PopupScreen "Tank 6S Status" 480x272
   TextField "Text field_4" at 9,135 size 86x22; Text 'Pressure:'
   IOField "I/O field_1" at 148,130 size 90x25; FormatPattern s999.9; Unit  mBar
      ProcessValue <- "20_TANKS_IP_DATA_RIO_06_SECOND_TANK_TANKS_PRESS"
   TextField "Text field_5" at 9,169 size 113x22; Text 'Water Level:'
   IOField "I/O field_2" at 148,164 size 90x25; FormatPattern 999.9; Unit  %
      ProcessValue <- "20_TANKS_IP_DATA_RIO_06_SECOND_TANK_BWT_LEVEL"
   TextField "Text field_6" at 9,203 size 137x22; Text 'MBG Flow Rate:'
   IOField "I/O field_3" at 148,198 size 90x25; FormatPattern 999.9; Unit  m³/hr
      ProcessValue <- "20_TANKS_IP_DATA_RIO_06_SECOND_TANK_MBG_FLOW"
   TextField "Text field_7" at 9,237 size 135x22; Text 'USD Flow Rate:'
   IOField "I/O field_4" at 148,232 size 90x25; FormatPattern 999.9; Unit  m³/hr
      ProcessValue <- "20_TANKS_IP_DATA_RIO_06_SECOND_TANK_USD_FLOW"
   Button "Button_1" at 51,5 size 191x35; TextOff 'Starboard Tank 6 (6S)'
      on Release: function_efd93a16("Tank 6S Status", 0, 0, -1, 2, 1)
   TextField "Text field_1" at 6,90 size 109x25; Text 'TIME LEFT:'
   GraphicView "Graphic view_1" at 9,46 size 228x32; Picture "Tank Manually Disabled"
   GraphicIOField "Graphic I/O field_1" at 9,46 size 228x32; PictureList "Tank Process Stage_II"
      ProcessValue <- "2100_BTCS_CNTRL_DB_BTCS_STATE"
      Visibility <- "504_Tank Grouping_DB2020_GROUP of TANK 13"
   Button "Button_2" at 4,5 size 45x35; TextOff 'Text'; PictureOff "Graphic_286"
      on Click: function_efd93a16("Tank 6S Status", 0, 0, -1, -1, 1)
   IOField "I/O field_29" at 190,90 size 47x25; FormatPattern 99; Unit m
      ProcessValue <- "504_Tank Grouping_DB2020_Time Left Tank_Time Left m Tank 13"
   IOField "I/O field_8" at 147,90 size 42x25; FormatPattern 99; Unit h
      ProcessValue <- "504_Tank Grouping_DB2020_Time Left Tank_Time Left h Tank 13"
   IOField "I/O field_9" at 104,90 size 42x25; FormatPattern 99; Unit d
      ProcessValue <- "504_Tank Grouping_DB2020_Time Left Tank_Time Left d Tank 13"
   TextField "Text field_8" at 244,135 size 140x22; Text 'Water pH Level:'
   IOField "I/O field_5" at 384,130 size 90x25; FormatPattern 99.9
      ProcessValue <- "20_TANKS_IP_DATA_RIO_06_SECOND_TANK_BWT_PH"
   TextField "Text field_9" at 244,169 size 143x22; Text 'Water DO Level:'
   IOField "I/O field_6" at 384,164 size 90x25; FormatPattern 99.99; Unit  mg/l
      ProcessValue <- "20_TANKS_IP_DATA_RIO_06_SECOND_TANK_BWT_DO"
   TextField "Text field_10" at 244,203 size 174x22; Text 'Water Temperature:'
   IOField "I/O field_7" at 399,198 size 75x25; FormatPattern 999.9; Unit  °C
      ProcessValue <- "20_TANKS_IP_DATA_RIO_06_SECOND_TANK_BWT_TEMP"
   Group "Group" at 248,228 size 226x40
   Button "Button_5" at 248,228 size 226x40; TextOff 'Tank Shutdown Alarm'
      Visibility <- "2062_Warning_Data_Alarm Tank S6"
   Button "Button_6" at 248,228 size 226x40; TextOff 'No/Low Water Level'; Authorization "Operate"
      Visibility <- "LT421 6S  TANK LEVEL ALARM_ALARM L"

PopupScreen "Tank 6P Status" 480x272
   TextField "Text field_4" at 9,135 size 86x22; Text 'Pressure:'
   IOField "I/O field_1" at 147,130 size 90x25; FormatPattern s999.9; Unit  mBar
      ProcessValue <- "20_TANKS_IP_DATA_RIO_06_FIRST_TANK_TANKS_PRESS"
   TextField "Text field_5" at 9,169 size 113x22; Text 'Water Level:'
   IOField "I/O field_2" at 147,164 size 90x25; FormatPattern 999.9; Unit  %
      ProcessValue <- "20_TANKS_IP_DATA_RIO_06_FIRST_TANK_BWT_LEVEL"
   TextField "Text field_6" at 9,203 size 137x22; Text 'MBG Flow Rate:'
   IOField "I/O field_3" at 147,198 size 90x25; FormatPattern 999.9; Unit  m³/hr
      ProcessValue <- "20_TANKS_IP_DATA_RIO_06_FIRST_TANK_MBG_FLOW"
   TextField "Text field_7" at 9,237 size 135x22; Text 'USD Flow Rate:'
   IOField "I/O field_4" at 147,232 size 90x25; FormatPattern 999.9; Unit  m³/hr
      ProcessValue <- "20_TANKS_IP_DATA_RIO_06_FIRST_TANK_USD_FLOW"
   Button "Button_1" at 51,5 size 190x35; TextOff 'Port Tank 6 (6P)'
      on Release: function_efd93a16("Tank 6P Status", 0, 0, -1, 2, 1)
   TextField "Text field_1" at 5,90 size 109x25; Text 'TIME LEFT:'
   GraphicView "Graphic view_1" at 9,46 size 227x32; Picture "Tank Manually Disabled"
   GraphicIOField "Graphic I/O field_1" at 9,46 size 227x32; PictureList "Tank Process Stage_II"
      ProcessValue <- "2100_BTCS_CNTRL_DB_BTCS_STATE"
      Visibility <- "504_Tank Grouping_DB2020_GROUP of TANK 12"
   Button "Button_2" at 4,5 size 45x35; TextOff 'Text'; PictureOff "Graphic_286"
      on Click: function_efd93a16("Tank 6P Status", 0, 0, -1, -1, 1)
   IOField "I/O field_29" at 189,90 size 47x25; FormatPattern 99; Unit m
      ProcessValue <- "504_Tank Grouping_DB2020_Time Left Tank_Time Left m Tank 12"
   IOField "I/O field_8" at 146,90 size 42x25; FormatPattern 99; Unit h
      ProcessValue <- "504_Tank Grouping_DB2020_Time Left Tank_Time Left h Tank 12"
   IOField "I/O field_9" at 103,90 size 42x25; FormatPattern 99; Unit d
      ProcessValue <- "504_Tank Grouping_DB2020_Time Left Tank_Time Left d Tank 12"
   TextField "Text field_8" at 242,135 size 140x22; Text 'Water pH Level:'
   IOField "I/O field_5" at 381,130 size 90x25; FormatPattern 99.9
      ProcessValue <- "20_TANKS_IP_DATA_RIO_06_FIRST_TANK_BWT_PH"
   TextField "Text field_9" at 242,169 size 143x22; Text 'Water DO Level:'
   IOField "I/O field_6" at 381,164 size 90x25; FormatPattern 99.99; Unit  mg/l
      ProcessValue <- "20_TANKS_IP_DATA_RIO_06_FIRST_TANK_BWT_DO"
   TextField "Text field_10" at 242,203 size 174x22; Text 'Water Temperature:'
   IOField "I/O field_7" at 396,198 size 75x25; FormatPattern 999.9; Unit  °C
      ProcessValue <- "20_TANKS_IP_DATA_RIO_06_FIRST_TANK_BWT_TEMP"
   Group "Group" at 245,227 size 226x40
   Button "Button_5" at 245,227 size 226x40; TextOff 'Tank Shutdown Alarm'
      Visibility <- "2062_Warning_Data_Alarm Tank P6"
   Button "Button_6" at 245,227 size 226x40; TextOff 'No/Low Water Level'; Authorization "Operate"
      Visibility <- "LT422 6P  TANK LEVEL ALARM_ALARM L"

PopupScreen "Tank AP Status" 480x272
   TextField "Text field_4" at 9,135 size 86x22; Text 'Pressure:'
   IOField "I/O field_1" at 147,130 size 90x25; FormatPattern s999.9; Unit  mBar
      ProcessValue <- "20_TANKS_IP_DATA_RIO_07_FIRST_TANK_TANKS_PRESS"
   TextField "Text field_5" at 9,169 size 113x22; Text 'Water Level:'
   IOField "I/O field_2" at 147,164 size 90x25; FormatPattern 999.9; Unit  %
      ProcessValue <- "20_TANKS_IP_DATA_RIO_07_FIRST_TANK_BWT_LEVEL"
   TextField "Text field_6" at 9,203 size 137x22; Text 'MBG Flow Rate:'
   IOField "I/O field_3" at 147,198 size 90x25; FormatPattern 999.9; Unit  m³/hr
      ProcessValue <- "20_TANKS_IP_DATA_RIO_07_FIRST_TANK_MBG_FLOW"
   TextField "Text field_7" at 9,237 size 135x22; Text 'USD Flow Rate:'
   IOField "I/O field_4" at 147,232 size 90x25; FormatPattern 999.9; Unit  m³/hr
      ProcessValue <- "20_TANKS_IP_DATA_RIO_07_FIRST_TANK_USD_FLOW"
   Button "Button_1" at 51,5 size 189x35; TextOff 'Aft Peak Tank (APT)'
      on Release: function_efd93a16("Tank AP Status", 0, 0, -1, 2, 1)
   TextField "Text field_1" at 5,90 size 109x25; Text 'TIME LEFT:'
   GraphicView "Graphic view_1" at 9,46 size 227x32; Picture "Tank Manually Disabled"
   GraphicIOField "Graphic I/O field_1" at 9,46 size 227x32; PictureList "Tank Process Stage_II"
      ProcessValue <- "2100_BTCS_CNTRL_DB_BTCS_STATE"
      Visibility <- "504_Tank Grouping_DB2020_GROUP of TANK 14"
   Button "Button_2" at 4,5 size 45x35; TextOff 'Text'; PictureOff "Graphic_286"
      on Click: function_efd93a16("Tank AP Status", 0, 0, -1, -1, 1)
   IOField "I/O field_29" at 189,90 size 47x25; FormatPattern 99; Unit m
      ProcessValue <- "504_Tank Grouping_DB2020_Time Left Tank_Time Left m Tank 14"
   IOField "I/O field_8" at 146,90 size 42x25; FormatPattern 99; Unit h
      ProcessValue <- "504_Tank Grouping_DB2020_Time Left Tank_Time Left h Tank 14"
   IOField "I/O field_9" at 103,90 size 42x25; FormatPattern 99; Unit d
      ProcessValue <- "504_Tank Grouping_DB2020_Time Left Tank_Time Left d Tank 14"
   TextField "Text field_8" at 245,135 size 140x22; Text 'Water pH Level:'
   IOField "I/O field_5" at 384,130 size 90x25; FormatPattern 99.9
      ProcessValue <- "20_TANKS_IP_DATA_RIO_07_FIRST_TANK_BWT_PH"
   TextField "Text field_9" at 245,169 size 143x22; Text 'Water DO Level:'
   IOField "I/O field_6" at 384,164 size 90x25; FormatPattern 99.99; Unit  mg/l
      ProcessValue <- "20_TANKS_IP_DATA_RIO_07_FIRST_TANK_BWT_DO"
   TextField "Text field_10" at 245,203 size 174x22; Text 'Water Temperature:'
   IOField "I/O field_7" at 399,198 size 75x25; FormatPattern 999.9; Unit  °C
      ProcessValue <- "20_TANKS_IP_DATA_RIO_07_FIRST_TANK_BWT_TEMP"
   Group "Group" at 246,228 size 228x40
   Button "Button_5" at 246,228 size 228x40; TextOff 'Tank Shutdown Alarm'
      Visibility <- "2062_Warning_Data_Alarm Tank APT"
   Button "Button_6" at 246,228 size 228x40; TextOff 'No/Low Water Level'; Authorization "Operate"
      Visibility <- "LT422 APT  TANK LEVEL ALARM_ALARM L"

PopupScreen "Tank FP Status" 480x272
   TextField "Text field_1" at 5,85 size 109x25; Text 'TIME LEFT:'
   TextField "Text field_4" at 9,130 size 86x22; Text 'Pressure:'
   IOField "I/O field_1" at 142,125 size 90x25; FormatPattern s999.9; Unit  mBar
      ProcessValue <- "20_TANKS_IP_DATA_RIO_01_FIRST_TANK_TANKS_PRESS"
   TextField "Text field_5" at 9,164 size 113x22; Text 'Water Level:'
   IOField "I/O field_2" at 142,159 size 90x25; FormatPattern 999.9; Unit  %
      ProcessValue <- "20_TANKS_IP_DATA_RIO_01_FIRST_TANK_BWT_LEVEL"
   TextField "Text field_6" at 9,198 size 137x22; Text 'MBG Flow Rate:'
   IOField "I/O field_3" at 142,193 size 90x25; FormatPattern 999.9; Unit  m³/hr
      ProcessValue <- "20_TANKS_IP_DATA_RIO_01_FIRST_TANK_MBG_FLOW"
   TextField "Text field_7" at 9,232 size 135x22; Text 'USD Flow Rate:'
   IOField "I/O field_4" at 142,227 size 90x25; FormatPattern 999.9; Unit  m³/hr
      ProcessValue <- "20_TANKS_IP_DATA_RIO_01_FIRST_TANK_USD_FLOW"
   TextField "Text field_8" at 243,129 size 140x22; Text 'Water pH Level:'
   IOField "I/O field_5" at 380,124 size 90x25; FormatPattern 99.9
      ProcessValue <- "20_TANKS_IP_DATA_RIO_01_FIRST_TANK_BWT_PH"
   TextField "Text field_9" at 243,163 size 143x22; Text 'Water DO Level:'
   IOField "I/O field_6" at 380,158 size 90x25; FormatPattern 99.99; Unit  mg/l
      ProcessValue <- "20_TANKS_IP_DATA_RIO_01_FIRST_TANK_BWT_DO"
   TextField "Text field_10" at 240,197 size 174x22; Text 'Water Temperature:'
   IOField "I/O field_7" at 395,192 size 75x25; FormatPattern 999.9; Unit  °C
      ProcessValue <- "20_TANKS_IP_DATA_RIO_01_FIRST_TANK_BWT_TEMP"
   IOField "I/O field_29" at 188,85 size 47x25; FormatPattern 99; Unit m
      ProcessValue <- "504_Tank Grouping_DB2020_Time Left Tank_Time Left m Tank 1"
   GraphicView "Graphic view_1" at 9,41 size 227x32; Picture "Tank Manually Disabled"
   Button "Button_1" at 49,1 size 192x35; TextOff 'Fore Peak Tank (FPT)'
   GraphicIOField "Graphic I/O field_1" at 9,41 size 227x32; PictureList "Tank Process Stage_II"
      ProcessValue <- "2100_BTCS_CNTRL_DB_BTCS_STATE"
      Visibility <- "504_Tank Grouping_DB2020_GROUP of TANK 1"
   Button "Button_7" at 4,1 size 43x35; TextOff 'Text'; PictureOff "Graphic_286"
      on Click: function_efd93a16("Tank FP Status", 0, 0, -1, -1, 1)
   IOField "I/O field_8" at 145,85 size 42x25; FormatPattern 99; Unit h
      ProcessValue <- "504_Tank Grouping_DB2020_Time Left Tank_Time Left h Tank 1"
   IOField "I/O field_9" at 102,85 size 42x25; FormatPattern 99; Unit d
      ProcessValue <- "504_Tank Grouping_DB2020_Time Left Tank_Time Left d Tank 1"
   Group "Group" at 271,226 size 195x40
   Button "Button_5" at 271,226 size 195x40; TextOff 'Tank Shutdown Alarm'
      Visibility <- "2062_Warning_Data_Alarm Tank FPT"
      ProcessValue <- "2062_Warning_Data_Water Level Override FPT"
   Button "Button_6" at 271,226 size 195x40; TextOff 'No/Low Water Level'
      ProcessValue <- "2062_Warning_Data_Water Level Override FPT"
      Visibility <- "LT422 FPT  TANK LEVEL ALARM_ALARM L"

PopupScreen "Info" 400x272
   TextField "Text field_3" at 6,135 size 94x28; Text 'Contact:'
   TextField "Text field_5" at 5,113 size 161x25; Text 'September 2018'
   GraphicView "Logo" at 4,3 size 219x60; Picture "Logo of IGG HMI"
   TextField "Text field_8" at 6,159 size 270x46; Text 'Coldharbour Marine Limited United Kingdom'
   TextField "Text field_9" at 6,200 size 386x67; Text 'T: +44 (0) 1629 888386 F: +44 (0) 1629 888385 E: techsupport@coldharbourmarine.com'
   TextField "Text field_1" at 5,71 size 415x46; Text '2 Tanks Ballast Water Treatment System Automation Control Software, Version 6.21'

SlideinScreen "GraphX_Slidein_Left" 158x272
   TextField "Text field_1" at 0,19 size 132x10; Text 'Inert Gas Generator Control Software'
   TextField "Text field_2" at 0,27 size 44x10; Text 'Version 3.0'
   TextField "Text field_3" at 0,65 size 43x10; Text 'Created by'
   TextField "Text field_4" at 0,73 size 127x11; Text 'Martin Ashiedu CEng MIET'
   TextField "Text field_5" at 0,35 size 57x10; Text 'December 2015'
   TextField "Text field_6" at 0,81 size 117x11; Text 'Coldharbour Marine Ltd'
   TextField "Text field_7" at 0,89 size 72x11; Text 'December 2015'

SlideinScreen "GraphX_Slidein_Bottom" 480x90
   TrendView "Trend view_1" at 0,0 size 480x92

PopupScreen "Start Treatment" 470x220
   Group "Group" at -16,2 size 485x220
   Button "Button_1" at 1,2 size 468x220; TextOff 'Text'
   Button "Button_2" at 144,134 size 174x55; TextOff 'OK'
      on Release: ResetBit("2102_TIME_CALCS_DB_PRE-DWEL_Warning 2"); function_efd93a16("Start Treatment", 0, 0, -1, -1, 1)
   TextField "Text field_1" at -16,53 size 455x40; Text 'Treatment now required'

PopupScreen "SD Card overflow" 468x220
   Button "Button_1" at 0,0 size 468x220; TextOff 'Data Logging SD Card Memory Full'
      on Click: function_efd93a16("SD Card overflow", 0, 0, -1, -1, 1)
      on Press: ResetBit("Logging SD Card Overflow")

PopupScreen "Time Until Treatment Required" 468x220
   Button "Button_1" at 0,0 size 468x220; TextOff 'Text'
   Button "Button_2" at 123,134 size 200x55; TextOff 'OK'
      on Release: ResetBit("2102_TIME_CALCS_DB_PRE-DWEL_Warning 1")
   TextField "Text field_1" at -77,20 size 557x104; Text 'Treatment required to start in hours and minutes'
   IOField "I/O field_1" at 178,54 size 47x40; FormatPattern 99
      ProcessValue <- "Sequence Times_DB_Pre-Dwell Timer_Hours Left"
   IOField "I/O field_2" at 199,89 size 47x40; FormatPattern 99
      ProcessValue <- "Sequence Times_DB_Pre-Dwell Timer_Minutes Left"

PopupScreen "Treatment check / Daily Checks Completed" 468x220
   Button "Button_3" at 117,134 size 229x50; TextOff 'CONFIRM'
      on Release: function_efd93a16("Treatment check / Daily Checks Completed", 0, 0, 0, -1, 1)
      on Press: function_b14e0dd5("88_treatment_POP_UP_CNFRM", 0)
   TextField "Text field_1" at 14,5 size 432x106; Text 'Please confirm pre treatment check and daily checks are completed.'

PopupScreen "Treatment Cycle Completed" 468x220
   Button "Button_1" at 0,0 size 468x220; TextOff 'TREATMENT CYCLE COMPLETED'
      on Click: function_efd93a16("Treatment Cycle Completed", 0, 0, -1, -1, 1)

PopupScreen "Treatment Status" 300x248
   Button "HmiScreenItemData_40" at 0,0 size 300x29; TextOn 'Back'; TextOff 'Treatment Status'
      on Release: function_efd93a16("Treatment Status", 0, 0, -1, -1, 1)
   Button "HmiScreenItemData_9" at 17,34 size 220x30; TextOn 'Back'; TextOff 'Pre Dwell Time Completed'
      on Release: function_efd93a16("Treatment Status", 0, 0, -1, -1, 1)
   Button "HmiScreenItemData_17" at 17,94 size 220x30; TextOn 'Back'; TextOff 'De-Oxygenation Completed'
      on Release: function_efd93a16("Treatment Status", 0, 0, -1, -1, 1)
   Button "HmiScreenItemData_38" at 17,124 size 220x30; TextOn 'Back'; TextOff 'Dwell Time Completed'
      on Release: function_efd93a16("Treatment Status", 0, 0, -1, -1, 1)
   Button "HmiScreenItemData_39" at 17,184 size 220x30; TextOn 'Back'; TextOff 'Re-Oxygenation Completed'
      on Release: function_efd93a16("Treatment Status", 0, 0, -1, -1, 1)
   Button "HmiScreenItemData_41" at 18,215 size 220x30; TextOn 'Back'; TextOff 'Post Dwell Time Completed'
      on Release: function_efd93a16("Treatment Status", 0, 0, -1, -1, 1)
   Button "HmiScreenItemData_46" at 17,64 size 220x30; TextOn 'Back'; TextOff 'Inert Gas Transfer Active'
   Button "HmiScreenItemData_48" at 17,154 size 220x30; TextOn 'Back'; TextOff 'Ambient Air Transfer Active'
   Button "HmiScreenItemData_52" at 17,64 size 220x30; TextOn 'Back'; TextOff 'IG Transfer Completed'
      on Release: function_efd93a16("Treatment Status", 0, 0, -1, -1, 1)
   Button "HmiScreenItemData_53" at 17,154 size 220x30; TextOn 'Back'; TextOff 'Ambient Air Transfer Completed'
      on Release: function_efd93a16("Treatment Status", 0, 0, -1, -1, 1)
   Button "Button_2" at 0,0 size 34x29; TextOff 'Text'; PictureOff "Graphic_286"
      on Click: function_efd93a16("Treatment Status", 0, 0, -1, -1, 1)
   Circle "Circle_23" at 254,38 size 24x24
      Appearance <- "2110_BTCS_CNTRL_DB_BTCS_STEP"
   Circle "Circle_24" at 254,67 size 24x24
      Appearance <- "100_GCU_AUTO_SEQ_DB_CRNT_STEP"
   Circle "Circle_25" at 254,97 size 24x24
      Appearance <- "2110_BTCS_CNTRL_DB_BTCS_STEP"
   Circle "Circle_26" at 254,127 size 24x24
      Appearance <- "2110_BTCS_CNTRL_DB_BTCS_STEP"
   Circle "Circle_27" at 254,157 size 24x24
      Appearance <- "100_GCU_AUTO_SEQ_DB_CRNT_STEP"
   Circle "Circle_28" at 254,187 size 24x24
      Appearance <- "2110_BTCS_CNTRL_DB_BTCS_STEP"
   Circle "Circle_29" at 254,217 size 24x24
      Appearance <- "2110_BTCS_CNTRL_DB_BTCS_STEP"

PopupScreen "Time Until GCU Start Required" 468x220
   Button "Button_1" at 0,0 size 468x220; TextOff 'Text'
   Button "Button_2" at 125,172 size 200x44; TextOff 'OK'; Authorization "Operate"
      on Release: function_efd93a16("Time Until GCU Start Required", 0, 0, -1, -1, 1); ActivateScreen("GCU Plant", 0)
   TextField "Text field_1" at -12,-3 size 490x112; Text 'Instalation Start Confirmation Required in hours for Re-Ox Stage'
   TextField "Text field_2" at 63,100 size 327x76; Text 'Please Make Sure the Energy and Water Supply are Present and Sufficient'
   IOField "I/O field_1" at 233,25 size 104x52; FormatPattern 99
      ProcessValue <- "Sequence Times_DB_Dwell Timer_Hours Left"

PopupScreen "Start GCU for Re-Ox" 468x220
   Button "Button_1" at 0,0 size 468x220; TextOff 'Text'
   Button "Button_2" at 133,154 size 200x55; TextOff 'OK'; Authorization "Operate"
      on Release: function_efd93a16("Start GCU for Re-Ox", 0, 0, -1, -1, 1); ActivateScreen("GCU Plant", 0)
   TextField "Text field_1" at -11,8 size 490x76; Text 'Instalation Start Confirmation Required for Re-Ox Stage'
   TextField "Text field_2" at 73,80 size 327x76; Text 'Please Make Sure the Energy and Water Supply are Present and Sufficient'

VB script "BWT_Warning"
   If SmartTags("BWT Mode Warning") Then
   	efd93a16-2665-4b85-bcb9-25eddcb7b6f4 BWT Mode Warning,275,250,$3$hmiOn$,$3$hmiTop$,$3$hmiMedium$
   'ElseIf Not SmartTags("BWT Mode Warning") Then
   '	ShowPopupScreen"BWT Mode Warning",0,0,hmiOff,hmiAnimationOff,hmiMedium
   End If

VB script "Report_Test"
   f41c6f6c-971d-4734-9362-16d81ac70597 Current User
   e1ab61de-e5a2-437b-97c4-abda991a3a2e user_group
   
   
   
   	
   	
   'Tip:
   ' 1. Use the <CTRL+SPACE> or <CTRL+I> shortcut to open a list of all objects and functions
   ' 2. Write the code using the HMI Runtime object.
   '  Example: HmiRuntime.Screens("Screen_1").
   ' 3. Use the <CTRL+J> shortcut to create an object reference.
   'Write the code as of this position:

VB script "SD_Card_Overflow"
   If SmartTags("Logging SD Card Overflow") Then 
   	efd93a16-2665-4b85-bcb9-25eddcb7b6f4 SD Card overflow,275,250,$3$hmiOn$,$3$hmiBottom$,$3$hmiMedium$
   ElseIf Not SmartTags("Logging SD Card Overflow") Then
   	efd93a16-2665-4b85-bcb9-25eddcb7b6f4SD Card overflow,0,0,$3$hmiOff$,$3$hmiAnimationOff$,$3$hmiMedium$
   End If

VB script "TitleUpdater"
   Dim title
   Set title = HmiRuntime.ActiveScreen.ScreenItems("Screen title")
   title.Text = HmiRuntime.ActiveScreen.ObjectName

VB script "TreatmentCycleCompleted"
   If SmartTags("Treatment Runs Completed") Then
   	efd93a16-2665-4b85-bcb9-25eddcb7b6f4 Treatment Cycle Completed,275,250,$3$hmiOn$,$3$hmiBottom$,$3$hmiMedium$
   'ElseIf Not SmartTags("Treatment Runs Completed") Then
   '	ShowPopupScreen"Treatment Cycle Completed",0,0,hmiOff,hmiAnimationOff,hmiMedium
   End If

VB script "TreatmentdDailyChecks"
   If SmartTags("88_treatment_POP_UP") Then
   	efd93a16-2665-4b85-bcb9-25eddcb7b6f4 Treatment check / Daily Checks Completed,275,250,$3$hmiOn$,$3$hmiBottom$,$3$hmiMedium$
   End If

VB script "User_Change"
   f41c6f6c-971d-4734-9362-16d81ac70597 Current User
   e1ab61de-e5a2-437b-97c4-abda991a3a2e user_group
   
   'Tip:
   ' 1. Use the <CTRL+SPACE> or <CTRL+I> shortcut to open a list of all objects and functions
   ' 2. Write the code using the HMI Runtime object.
   '  Example: HmiRuntime.Screens("Screen_1").
   ' 3. Use the <CTRL+J> shortcut to create an object reference.
   'Write the code as of this position:

VB script "Buzzer"
   Dim Buzz
   If SmartTags("Shutdown Alarm") Then 
   	bec8f1e5-2ab1-45f6-ad91-1d37c469eb91Alarm.Alarms,0,0,$3$hmiOn$,$3$hmiBottom$,$3$hmiMedium$
   Set Buzz = HmiRuntime.ActiveScreen.ScreenItems("Alarm.Alarms.Media Player_1")
   Buzz = True
   
   
   
   
   'Tip:
   ' 1. Use the <CTRL+SPACE> or <CTRL+I> shortcut to open a list of all objects and functions
   ' 2. Write the code using the HMI Runtime object.
   '  Example: HmiRuntime.Screens("Screen_1").
   ' 3. Use the <CTRL+J> shortcut to create an object reference.
   'Write the code as of this position:

VB script "HeartBeatFunction"
   Dim TimerAux
   
   If SmartTags("BRIGE HMI HEART BEAT")=0 Then
   	b21d3eaf-4e31-425c-ad1a-ba4e4002cacc(BRIGE HMI HEART BEAT),1
   Else
   	b21d3eaf-4e31-425c-ad1a-ba4e4002cacc (BRIGE HMI HEART BEAT),0
   End If
   
   'Tip:
   ' 1. Use the <CTRL+SPACE> or <CTRL+I> shortcut to open a list of all objects and functions
   ' 2. Write the code using the HMI Runtime object.
   '  Example: HmiRuntime.Screens("Screen_1").
   ' 3. Use the <CTRL+J> shortcut to create an object reference.
   'Write the code as of this position:

VB script "ALARM_Present"
   If SmartTags("60_Alarm_Data_ALRM_PRSNT") Then
   	bec8f1e5-2ab1-45f6-ad91-1d37c469eb91 Alarms,0
   End If
   
   
   
   
   
   
   
   
   
   
   
   'Tip:
   ' 1. Use the <CTRL+SPACE> or <CTRL+I> shortcut to open a list of all objects and functions
   ' 2. Write the code using the HMI Runtime object.
   '  Example: HmiRuntime.Screens("Screen_1").
   ' 3. Use the <CTRL+J> shortcut to create an object reference.
   'Write the code as of this position:

VB script "TimeRemainingToRe_Ox"
   If SmartTags("Warn To Start GCU") Then
   	efd93a16-2665-4b85-bcb9-25eddcb7b6f4 Time Until GCU Start Required, 0, 0, $3$hmiOn$, $3$hmiBottom$, $3$hmiMedium$
   	ElseIf Not SmartTags("Warn To Start GCU") Then
   efd93a16-2665-4b85-bcb9-25eddcb7b6f4 Time Until GCU Start Required, 0, 0, $3$hmiOff$, $3$hmiOff$, $3$hmiMedium$
   End If

VB script "TimeRemainingToTreatment"
   If SmartTags("Warn To Start IGG") Then
   	efd93a16-2665-4b85-bcb9-25eddcb7b6f4 Time Until Treatment Required, 400, 200, $3$hmiOn$, $3$hmiBottom$, $3$hmiMedium$
   	ElseIf Not SmartTags("Warn To Start IGG") Then
   efd93a16-2665-4b85-bcb9-25eddcb7b6f4 Time Until Treatment Required, 0, 0, $3$hmiOff$, $3$hmiOff$, $3$hmiMedium$
   End If

VB script "TreatmentRequired"
   If SmartTags("Warn To Start IGG-Last") Then
   	efd93a16-2665-4b85-bcb9-25eddcb7b6f4 Start Treatment, 400, 200, $3$hmiOn$, $3$hmiBottom$, $3$hmiMedium$
   	ElseIf Not SmartTags("Warn To Start IGG-Last") Then
       efd93a16-2665-4b85-bcb9-25eddcb7b6f4 Start Treatment, 0, 0, $3$hmiOff$, $3$hmiOff$, $3$hmiMedium$
   End If

VB script "TreatmentRequired_GCU"
   If SmartTags("Warn To Start GCU-Last") Then
   	efd93a16-2665-4b85-bcb9-25eddcb7b6f4 Start GCU for Re-Ox, 0, 0, $3$hmiOn$, $3$hmiBottom$, $3$hmiMedium$
   	ElseIf Not SmartTags("Warn To Start GCU-Last") Then
   efd93a16-2665-4b85-bcb9-25eddcb7b6f4 Start GCU for Re-Ox, 0, 0, $3$hmiOff$, $3$hmiOff$, $3$hmiMedium$
   End If
*)